REGION Network 15: EM - Abort Command
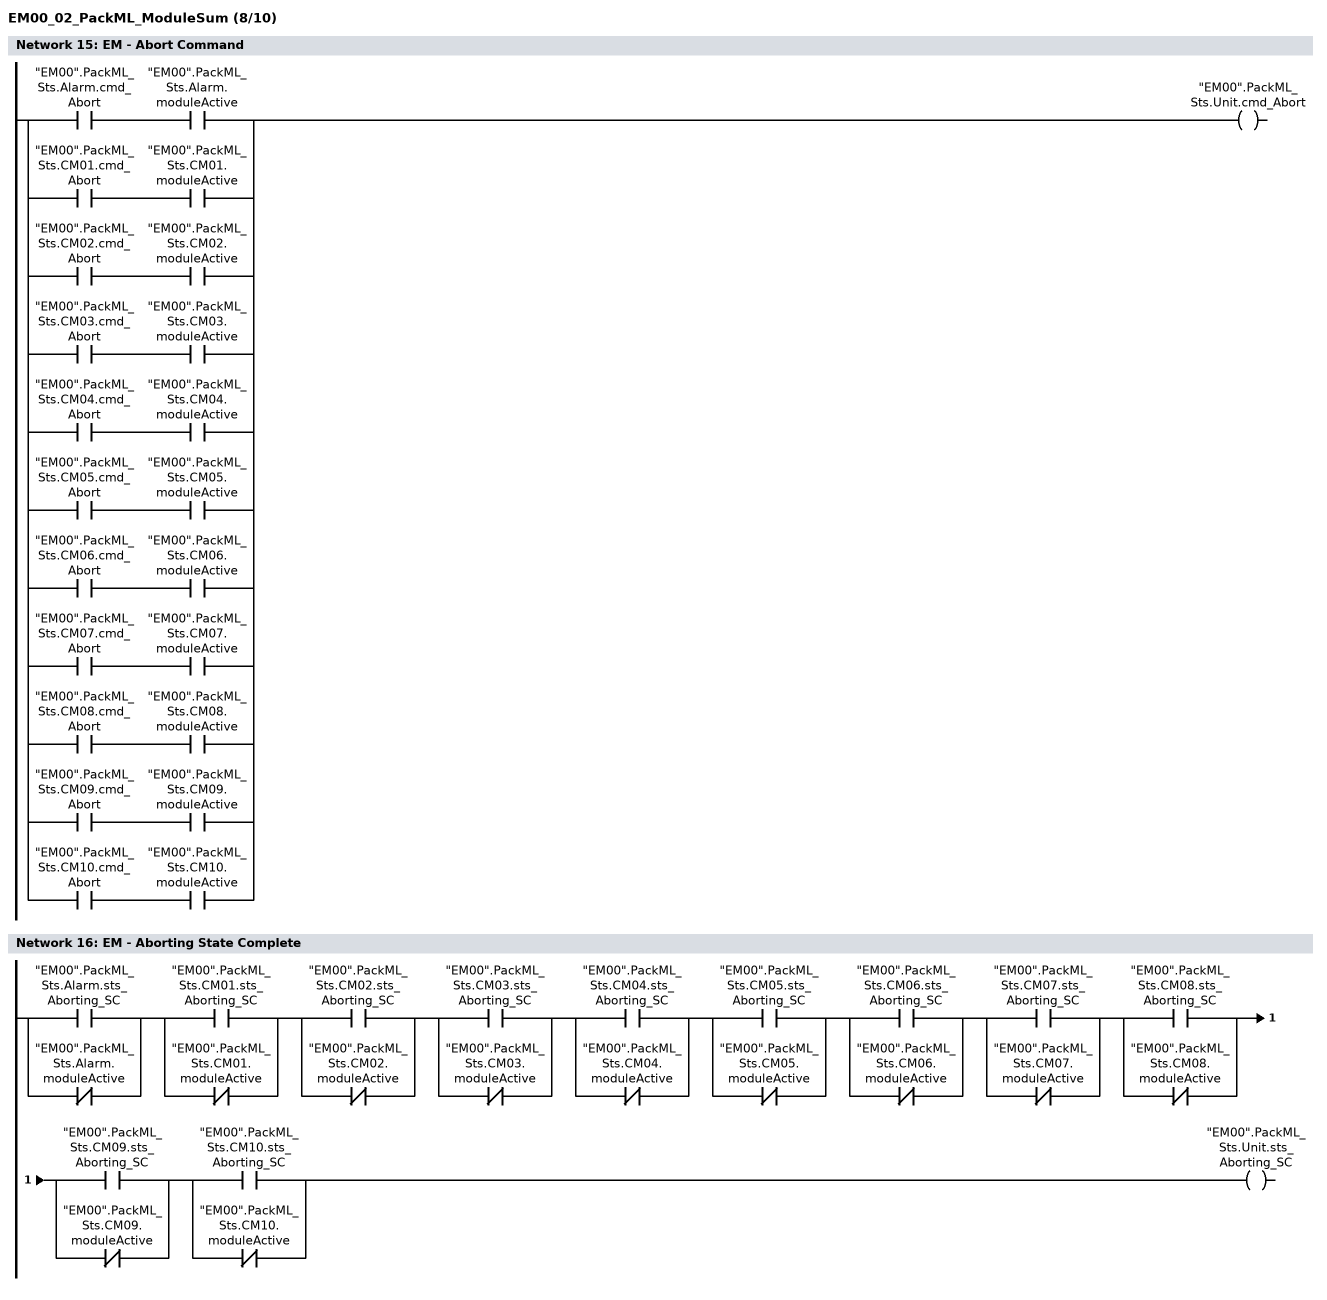
   RUNG wire#powerrail
      Contact( "EM00".PackML_Sts.Alarm.cmd_Abort )
      Contact( "EM00".PackML_Sts.Alarm.moduleActive )
      wire#w1
      Coil( "EM00".PackML_Sts.Unit.cmd_Abort )
   END_RUNG
   RUNG wire#powerrail
      Contact( "EM00".PackML_Sts.CM01.cmd_Abort )
      Contact( "EM00".PackML_Sts.CM01.moduleActive )
   END_RUNG wire#w1
   RUNG wire#powerrail
      Contact( "EM00".PackML_Sts.CM02.cmd_Abort )
      Contact( "EM00".PackML_Sts.CM02.moduleActive )
   END_RUNG wire#w1
   RUNG wire#powerrail
      Contact( "EM00".PackML_Sts.CM03.cmd_Abort )
      Contact( "EM00".PackML_Sts.CM03.moduleActive )
   END_RUNG wire#w1
   RUNG wire#powerrail
      Contact( "EM00".PackML_Sts.CM04.cmd_Abort )
      Contact( "EM00".PackML_Sts.CM04.moduleActive )
   END_RUNG wire#w1
   RUNG wire#powerrail
      Contact( "EM00".PackML_Sts.CM05.cmd_Abort )
      Contact( "EM00".PackML_Sts.CM05.moduleActive )
   END_RUNG wire#w1
   RUNG wire#powerrail
      Contact( "EM00".PackML_Sts.CM06.cmd_Abort )
      Contact( "EM00".PackML_Sts.CM06.moduleActive )
   END_RUNG wire#w1
   RUNG wire#powerrail
      Contact( "EM00".PackML_Sts.CM07.cmd_Abort )
      Contact( "EM00".PackML_Sts.CM07.moduleActive )
   END_RUNG wire#w1
   RUNG wire#powerrail
      Contact( "EM00".PackML_Sts.CM08.cmd_Abort )
      Contact( "EM00".PackML_Sts.CM08.moduleActive )
   END_RUNG wire#w1
   RUNG wire#powerrail
      Contact( "EM00".PackML_Sts.CM09.cmd_Abort )
      Contact( "EM00".PackML_Sts.CM09.moduleActive )
   END_RUNG wire#w1
   RUNG wire#powerrail
      Contact( "EM00".PackML_Sts.CM10.cmd_Abort )
      Contact( "EM00".PackML_Sts.CM10.moduleActive )
   END_RUNG wire#w1
   // the same network as SCL:
   "EM00".PackML_Sts.Unit.cmd_Abort := ("EM00".PackML_Sts.Alarm.cmd_Abort AND "EM00".PackML_Sts.Alarm.moduleActive) OR ("EM00".PackML_Sts.CM01.cmd_Abort AND "EM00".PackML_Sts.CM01.moduleActive) OR ("EM00".PackML_Sts.CM02.cmd_Abort AND "EM00".PackML_Sts.CM02.moduleActive) OR ("EM00".PackML_Sts.CM03.cmd_Abort AND "EM00".PackML_Sts.CM03.moduleActive) OR ("EM00".PackML_Sts.CM04.cmd_Abort AND "EM00".PackML_Sts.CM04.moduleActive) OR ("EM00".PackML_Sts.CM05.cmd_Abort AND "EM00".PackML_Sts.CM05.moduleActive) OR ("EM00".PackML_Sts.CM06.cmd_Abort AND "EM00".PackML_Sts.CM06.moduleActive) OR ("EM00".PackML_Sts.CM07.cmd_Abort AND "EM00".PackML_Sts.CM07.moduleActive) OR ("EM00".PackML_Sts.CM08.cmd_Abort AND "EM00".PackML_Sts.CM08.moduleActive) OR ("EM00".PackML_Sts.CM09.cmd_Abort AND "EM00".PackML_Sts.CM09.moduleActive) OR ("EM00".PackML_Sts.CM10.cmd_Abort AND "EM00".PackML_Sts.CM10.moduleActive);
END_REGION

REGION Network 16: EM - Aborting State Complete
   RUNG wire#powerrail
      Contact( "EM00".PackML_Sts.Alarm.sts_Aborting_SC )
      wire#w1
      Contact( "EM00".PackML_Sts.CM01.sts_Aborting_SC )
      wire#w2
      Contact( "EM00".PackML_Sts.CM02.sts_Aborting_SC )
      wire#w3
      Contact( "EM00".PackML_Sts.CM03.sts_Aborting_SC )
      wire#w4
      Contact( "EM00".PackML_Sts.CM04.sts_Aborting_SC )
      wire#w5
      Contact( "EM00".PackML_Sts.CM05.sts_Aborting_SC )
      wire#w6
      Contact( "EM00".PackML_Sts.CM06.sts_Aborting_SC )
      wire#w7
      Contact( "EM00".PackML_Sts.CM07.sts_Aborting_SC )
      wire#w8
      Contact( "EM00".PackML_Sts.CM08.sts_Aborting_SC )
      wire#w9
      Contact( "EM00".PackML_Sts.CM09.sts_Aborting_SC )
      wire#w10
      Contact( "EM00".PackML_Sts.CM10.sts_Aborting_SC )
      wire#w11
      Coil( "EM00".PackML_Sts.Unit.sts_Aborting_SC )
   END_RUNG
   RUNG wire#powerrail
      I_Contact( "EM00".PackML_Sts.Alarm.moduleActive )
   END_RUNG wire#w1
   RUNG wire#w1
      I_Contact( "EM00".PackML_Sts.CM01.moduleActive )
   END_RUNG wire#w2
   RUNG wire#w2
      I_Contact( "EM00".PackML_Sts.CM02.moduleActive )
   END_RUNG wire#w3
   RUNG wire#w3
      I_Contact( "EM00".PackML_Sts.CM03.moduleActive )
   END_RUNG wire#w4
   RUNG wire#w4
      I_Contact( "EM00".PackML_Sts.CM04.moduleActive )
   END_RUNG wire#w5
   RUNG wire#w5
      I_Contact( "EM00".PackML_Sts.CM05.moduleActive )
   END_RUNG wire#w6
   RUNG wire#w6
      I_Contact( "EM00".PackML_Sts.CM06.moduleActive )
   END_RUNG wire#w7
   RUNG wire#w7
      I_Contact( "EM00".PackML_Sts.CM07.moduleActive )
   END_RUNG wire#w8
   RUNG wire#w8
      I_Contact( "EM00".PackML_Sts.CM08.moduleActive )
   END_RUNG wire#w9
   RUNG wire#w9
      I_Contact( "EM00".PackML_Sts.CM09.moduleActive )
   END_RUNG wire#w10
   RUNG wire#w10
      I_Contact( "EM00".PackML_Sts.CM10.moduleActive )
   END_RUNG wire#w11
   // the same network as SCL:
   "EM00".PackML_Sts.Unit.sts_Aborting_SC := ("EM00".PackML_Sts.Alarm.sts_Aborting_SC OR NOT "EM00".PackML_Sts.Alarm.moduleActive) AND ("EM00".PackML_Sts.CM01.sts_Aborting_SC OR NOT "EM00".PackML_Sts.CM01.moduleActive) AND ("EM00".PackML_Sts.CM02.sts_Aborting_SC OR NOT "EM00".PackML_Sts.CM02.moduleActive) AND ("EM00".PackML_Sts.CM03.sts_Aborting_SC OR NOT "EM00".PackML_Sts.CM03.moduleActive) AND ("EM00".PackML_Sts.CM04.sts_Aborting_SC OR NOT "EM00".PackML_Sts.CM04.moduleActive) AND ("EM00".PackML_Sts.CM05.sts_Aborting_SC OR NOT "EM00".PackML_Sts.CM05.moduleActive) AND ("EM00".PackML_Sts.CM06.sts_Aborting_SC OR NOT "EM00".PackML_Sts.CM06.moduleActive) AND ("EM00".PackML_Sts.CM07.sts_Aborting_SC OR NOT "EM00".PackML_Sts.CM07.moduleActive) AND ("EM00".PackML_Sts.CM08.sts_Aborting_SC OR NOT "EM00".PackML_Sts.CM08.moduleActive) AND ("EM00".PackML_Sts.CM09.sts_Aborting_SC OR NOT "EM00".PackML_Sts.CM09.moduleActive) AND ("EM00".PackML_Sts.CM10.sts_Aborting_SC OR NOT "EM00".PackML_Sts.CM10.moduleActive);
END_REGION

REGION Network 17: EM - Clear Command
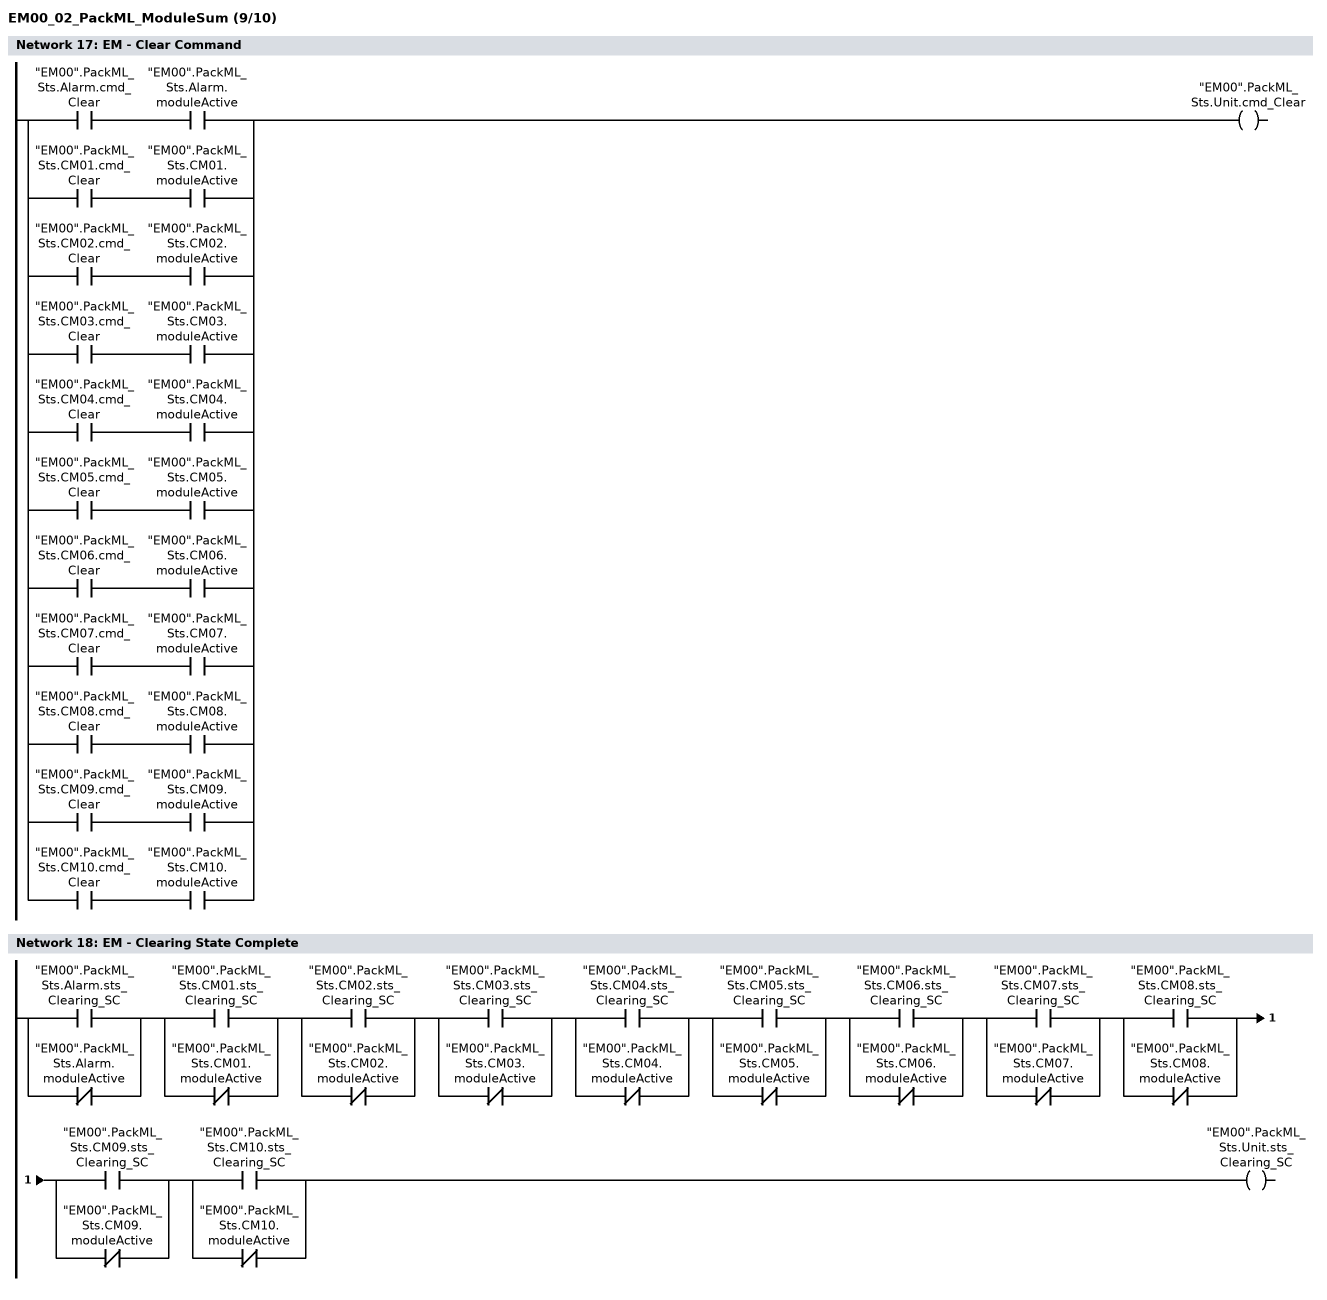
   RUNG wire#powerrail
      Contact( "EM00".PackML_Sts.Alarm.cmd_Clear )
      Contact( "EM00".PackML_Sts.Alarm.moduleActive )
      wire#w1
      Coil( "EM00".PackML_Sts.Unit.cmd_Clear )
   END_RUNG
   RUNG wire#powerrail
      Contact( "EM00".PackML_Sts.CM01.cmd_Clear )
      Contact( "EM00".PackML_Sts.CM01.moduleActive )
   END_RUNG wire#w1
   RUNG wire#powerrail
      Contact( "EM00".PackML_Sts.CM02.cmd_Clear )
      Contact( "EM00".PackML_Sts.CM02.moduleActive )
   END_RUNG wire#w1
   RUNG wire#powerrail
      Contact( "EM00".PackML_Sts.CM03.cmd_Clear )
      Contact( "EM00".PackML_Sts.CM03.moduleActive )
   END_RUNG wire#w1
   RUNG wire#powerrail
      Contact( "EM00".PackML_Sts.CM04.cmd_Clear )
      Contact( "EM00".PackML_Sts.CM04.moduleActive )
   END_RUNG wire#w1
   RUNG wire#powerrail
      Contact( "EM00".PackML_Sts.CM05.cmd_Clear )
      Contact( "EM00".PackML_Sts.CM05.moduleActive )
   END_RUNG wire#w1
   RUNG wire#powerrail
      Contact( "EM00".PackML_Sts.CM06.cmd_Clear )
      Contact( "EM00".PackML_Sts.CM06.moduleActive )
   END_RUNG wire#w1
   RUNG wire#powerrail
      Contact( "EM00".PackML_Sts.CM07.cmd_Clear )
      Contact( "EM00".PackML_Sts.CM07.moduleActive )
   END_RUNG wire#w1
   RUNG wire#powerrail
      Contact( "EM00".PackML_Sts.CM08.cmd_Clear )
      Contact( "EM00".PackML_Sts.CM08.moduleActive )
   END_RUNG wire#w1
   RUNG wire#powerrail
      Contact( "EM00".PackML_Sts.CM09.cmd_Clear )
      Contact( "EM00".PackML_Sts.CM09.moduleActive )
   END_RUNG wire#w1
   RUNG wire#powerrail
      Contact( "EM00".PackML_Sts.CM10.cmd_Clear )
      Contact( "EM00".PackML_Sts.CM10.moduleActive )
   END_RUNG wire#w1
   // the same network as SCL:
   "EM00".PackML_Sts.Unit.cmd_Clear := ("EM00".PackML_Sts.Alarm.cmd_Clear AND "EM00".PackML_Sts.Alarm.moduleActive) OR ("EM00".PackML_Sts.CM01.cmd_Clear AND "EM00".PackML_Sts.CM01.moduleActive) OR ("EM00".PackML_Sts.CM02.cmd_Clear AND "EM00".PackML_Sts.CM02.moduleActive) OR ("EM00".PackML_Sts.CM03.cmd_Clear AND "EM00".PackML_Sts.CM03.moduleActive) OR ("EM00".PackML_Sts.CM04.cmd_Clear AND "EM00".PackML_Sts.CM04.moduleActive) OR ("EM00".PackML_Sts.CM05.cmd_Clear AND "EM00".PackML_Sts.CM05.moduleActive) OR ("EM00".PackML_Sts.CM06.cmd_Clear AND "EM00".PackML_Sts.CM06.moduleActive) OR ("EM00".PackML_Sts.CM07.cmd_Clear AND "EM00".PackML_Sts.CM07.moduleActive) OR ("EM00".PackML_Sts.CM08.cmd_Clear AND "EM00".PackML_Sts.CM08.moduleActive) OR ("EM00".PackML_Sts.CM09.cmd_Clear AND "EM00".PackML_Sts.CM09.moduleActive) OR ("EM00".PackML_Sts.CM10.cmd_Clear AND "EM00".PackML_Sts.CM10.moduleActive);
END_REGION

REGION Network 18: EM - Clearing State Complete
   RUNG wire#powerrail
      Contact( "EM00".PackML_Sts.Alarm.sts_Clearing_SC )
      wire#w1
      Contact( "EM00".PackML_Sts.CM01.sts_Clearing_SC )
      wire#w2
      Contact( "EM00".PackML_Sts.CM02.sts_Clearing_SC )
      wire#w3
      Contact( "EM00".PackML_Sts.CM03.sts_Clearing_SC )
      wire#w4
      Contact( "EM00".PackML_Sts.CM04.sts_Clearing_SC )
      wire#w5
      Contact( "EM00".PackML_Sts.CM05.sts_Clearing_SC )
      wire#w6
      Contact( "EM00".PackML_Sts.CM06.sts_Clearing_SC )
      wire#w7
      Contact( "EM00".PackML_Sts.CM07.sts_Clearing_SC )
      wire#w8
      Contact( "EM00".PackML_Sts.CM08.sts_Clearing_SC )
      wire#w9
      Contact( "EM00".PackML_Sts.CM09.sts_Clearing_SC )
      wire#w10
      Contact( "EM00".PackML_Sts.CM10.sts_Clearing_SC )
      wire#w11
      Coil( "EM00".PackML_Sts.Unit.sts_Clearing_SC )
   END_RUNG
   RUNG wire#powerrail
      I_Contact( "EM00".PackML_Sts.Alarm.moduleActive )
   END_RUNG wire#w1
   RUNG wire#w1
      I_Contact( "EM00".PackML_Sts.CM01.moduleActive )
   END_RUNG wire#w2
   RUNG wire#w2
      I_Contact( "EM00".PackML_Sts.CM02.moduleActive )
   END_RUNG wire#w3
   RUNG wire#w3
      I_Contact( "EM00".PackML_Sts.CM03.moduleActive )
   END_RUNG wire#w4
   RUNG wire#w4
      I_Contact( "EM00".PackML_Sts.CM04.moduleActive )
   END_RUNG wire#w5
   RUNG wire#w5
      I_Contact( "EM00".PackML_Sts.CM05.moduleActive )
   END_RUNG wire#w6
   RUNG wire#w6
      I_Contact( "EM00".PackML_Sts.CM06.moduleActive )
   END_RUNG wire#w7
   RUNG wire#w7
      I_Contact( "EM00".PackML_Sts.CM07.moduleActive )
   END_RUNG wire#w8
   RUNG wire#w8
      I_Contact( "EM00".PackML_Sts.CM08.moduleActive )
   END_RUNG wire#w9
   RUNG wire#w9
      I_Contact( "EM00".PackML_Sts.CM09.moduleActive )
   END_RUNG wire#w10
   RUNG wire#w10
      I_Contact( "EM00".PackML_Sts.CM10.moduleActive )
   END_RUNG wire#w11
   // the same network as SCL:
   "EM00".PackML_Sts.Unit.sts_Clearing_SC := ("EM00".PackML_Sts.Alarm.sts_Clearing_SC OR NOT "EM00".PackML_Sts.Alarm.moduleActive) AND ("EM00".PackML_Sts.CM01.sts_Clearing_SC OR NOT "EM00".PackML_Sts.CM01.moduleActive) AND ("EM00".PackML_Sts.CM02.sts_Clearing_SC OR NOT "EM00".PackML_Sts.CM02.moduleActive) AND ("EM00".PackML_Sts.CM03.sts_Clearing_SC OR NOT "EM00".PackML_Sts.CM03.moduleActive) AND ("EM00".PackML_Sts.CM04.sts_Clearing_SC OR NOT "EM00".PackML_Sts.CM04.moduleActive) AND ("EM00".PackML_Sts.CM05.sts_Clearing_SC OR NOT "EM00".PackML_Sts.CM05.moduleActive) AND ("EM00".PackML_Sts.CM06.sts_Clearing_SC OR NOT "EM00".PackML_Sts.CM06.moduleActive) AND ("EM00".PackML_Sts.CM07.sts_Clearing_SC OR NOT "EM00".PackML_Sts.CM07.moduleActive) AND ("EM00".PackML_Sts.CM08.sts_Clearing_SC OR NOT "EM00".PackML_Sts.CM08.moduleActive) AND ("EM00".PackML_Sts.CM09.sts_Clearing_SC OR NOT "EM00".PackML_Sts.CM09.moduleActive) AND ("EM00".PackML_Sts.CM10.sts_Clearing_SC OR NOT "EM00".PackML_Sts.CM10.moduleActive);
END_REGION

REGION Network 19: EM - Execute State Complete
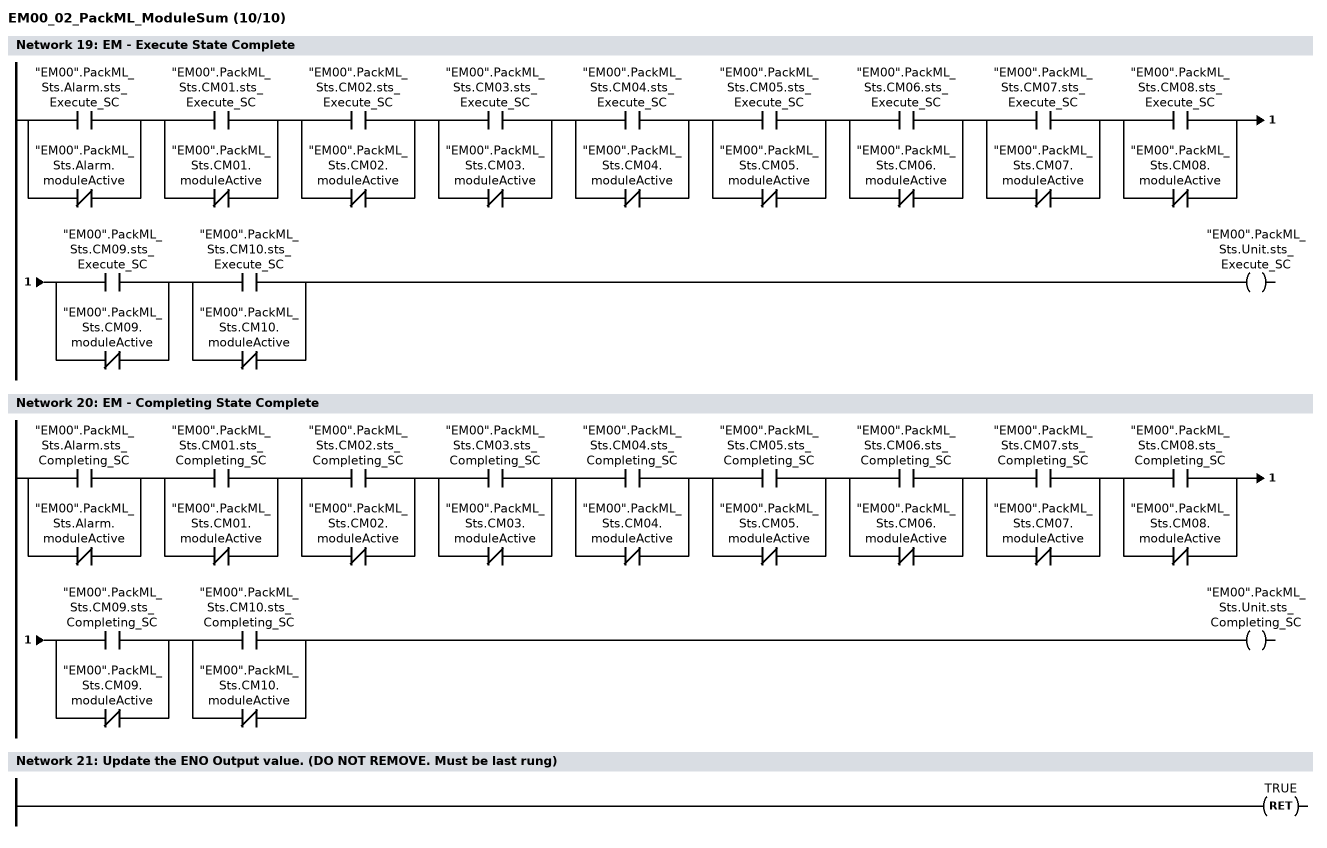
   RUNG wire#powerrail
      Contact( "EM00".PackML_Sts.Alarm.sts_Execute_SC )
      wire#w1
      Contact( "EM00".PackML_Sts.CM01.sts_Execute_SC )
      wire#w2
      Contact( "EM00".PackML_Sts.CM02.sts_Execute_SC )
      wire#w3
      Contact( "EM00".PackML_Sts.CM03.sts_Execute_SC )
      wire#w4
      Contact( "EM00".PackML_Sts.CM04.sts_Execute_SC )
      wire#w5
      Contact( "EM00".PackML_Sts.CM05.sts_Execute_SC )
      wire#w6
      Contact( "EM00".PackML_Sts.CM06.sts_Execute_SC )
      wire#w7
      Contact( "EM00".PackML_Sts.CM07.sts_Execute_SC )
      wire#w8
      Contact( "EM00".PackML_Sts.CM08.sts_Execute_SC )
      wire#w9
      Contact( "EM00".PackML_Sts.CM09.sts_Execute_SC )
      wire#w10
      Contact( "EM00".PackML_Sts.CM10.sts_Execute_SC )
      wire#w11
      Coil( "EM00".PackML_Sts.Unit.sts_Execute_SC )
   END_RUNG
   RUNG wire#powerrail
      I_Contact( "EM00".PackML_Sts.Alarm.moduleActive )
   END_RUNG wire#w1
   RUNG wire#w1
      I_Contact( "EM00".PackML_Sts.CM01.moduleActive )
   END_RUNG wire#w2
   RUNG wire#w2
      I_Contact( "EM00".PackML_Sts.CM02.moduleActive )
   END_RUNG wire#w3
   RUNG wire#w3
      I_Contact( "EM00".PackML_Sts.CM03.moduleActive )
   END_RUNG wire#w4
   RUNG wire#w4
      I_Contact( "EM00".PackML_Sts.CM04.moduleActive )
   END_RUNG wire#w5
   RUNG wire#w5
      I_Contact( "EM00".PackML_Sts.CM05.moduleActive )
   END_RUNG wire#w6
   RUNG wire#w6
      I_Contact( "EM00".PackML_Sts.CM06.moduleActive )
   END_RUNG wire#w7
   RUNG wire#w7
      I_Contact( "EM00".PackML_Sts.CM07.moduleActive )
   END_RUNG wire#w8
   RUNG wire#w8
      I_Contact( "EM00".PackML_Sts.CM08.moduleActive )
   END_RUNG wire#w9
   RUNG wire#w9
      I_Contact( "EM00".PackML_Sts.CM09.moduleActive )
   END_RUNG wire#w10
   RUNG wire#w10
      I_Contact( "EM00".PackML_Sts.CM10.moduleActive )
   END_RUNG wire#w11
   // the same network as SCL:
   "EM00".PackML_Sts.Unit.sts_Execute_SC := ("EM00".PackML_Sts.Alarm.sts_Execute_SC OR NOT "EM00".PackML_Sts.Alarm.moduleActive) AND ("EM00".PackML_Sts.CM01.sts_Execute_SC OR NOT "EM00".PackML_Sts.CM01.moduleActive) AND ("EM00".PackML_Sts.CM02.sts_Execute_SC OR NOT "EM00".PackML_Sts.CM02.moduleActive) AND ("EM00".PackML_Sts.CM03.sts_Execute_SC OR NOT "EM00".PackML_Sts.CM03.moduleActive) AND ("EM00".PackML_Sts.CM04.sts_Execute_SC OR NOT "EM00".PackML_Sts.CM04.moduleActive) AND ("EM00".PackML_Sts.CM05.sts_Execute_SC OR NOT "EM00".PackML_Sts.CM05.moduleActive) AND ("EM00".PackML_Sts.CM06.sts_Execute_SC OR NOT "EM00".PackML_Sts.CM06.moduleActive) AND ("EM00".PackML_Sts.CM07.sts_Execute_SC OR NOT "EM00".PackML_Sts.CM07.moduleActive) AND ("EM00".PackML_Sts.CM08.sts_Execute_SC OR NOT "EM00".PackML_Sts.CM08.moduleActive) AND ("EM00".PackML_Sts.CM09.sts_Execute_SC OR NOT "EM00".PackML_Sts.CM09.moduleActive) AND ("EM00".PackML_Sts.CM10.sts_Execute_SC OR NOT "EM00".PackML_Sts.CM10.moduleActive);
END_REGION

REGION Network 20: EM - Completing State Complete
   RUNG wire#powerrail
      Contact( "EM00".PackML_Sts.Alarm.sts_Completing_SC )
      wire#w1
      Contact( "EM00".PackML_Sts.CM01.sts_Completing_SC )
      wire#w2
      Contact( "EM00".PackML_Sts.CM02.sts_Completing_SC )
      wire#w3
      Contact( "EM00".PackML_Sts.CM03.sts_Completing_SC )
      wire#w4
      Contact( "EM00".PackML_Sts.CM04.sts_Completing_SC )
      wire#w5
      Contact( "EM00".PackML_Sts.CM05.sts_Completing_SC )
      wire#w6
      Contact( "EM00".PackML_Sts.CM06.sts_Completing_SC )
      wire#w7
      Contact( "EM00".PackML_Sts.CM07.sts_Completing_SC )
      wire#w8
      Contact( "EM00".PackML_Sts.CM08.sts_Completing_SC )
      wire#w9
      Contact( "EM00".PackML_Sts.CM09.sts_Completing_SC )
      wire#w10
      Contact( "EM00".PackML_Sts.CM10.sts_Completing_SC )
      wire#w11
      Coil( "EM00".PackML_Sts.Unit.sts_Completing_SC )
   END_RUNG
   RUNG wire#powerrail
      I_Contact( "EM00".PackML_Sts.Alarm.moduleActive )
   END_RUNG wire#w1
   RUNG wire#w1
      I_Contact( "EM00".PackML_Sts.CM01.moduleActive )
   END_RUNG wire#w2
   RUNG wire#w2
      I_Contact( "EM00".PackML_Sts.CM02.moduleActive )
   END_RUNG wire#w3
   RUNG wire#w3
      I_Contact( "EM00".PackML_Sts.CM03.moduleActive )
   END_RUNG wire#w4
   RUNG wire#w4
      I_Contact( "EM00".PackML_Sts.CM04.moduleActive )
   END_RUNG wire#w5
   RUNG wire#w5
      I_Contact( "EM00".PackML_Sts.CM05.moduleActive )
   END_RUNG wire#w6
   RUNG wire#w6
      I_Contact( "EM00".PackML_Sts.CM06.moduleActive )
   END_RUNG wire#w7
   RUNG wire#w7
      I_Contact( "EM00".PackML_Sts.CM07.moduleActive )
   END_RUNG wire#w8
   RUNG wire#w8
      I_Contact( "EM00".PackML_Sts.CM08.moduleActive )
   END_RUNG wire#w9
   RUNG wire#w9
      I_Contact( "EM00".PackML_Sts.CM09.moduleActive )
   END_RUNG wire#w10
   RUNG wire#w10
      I_Contact( "EM00".PackML_Sts.CM10.moduleActive )
   END_RUNG wire#w11
   // the same network as SCL:
   "EM00".PackML_Sts.Unit.sts_Completing_SC := ("EM00".PackML_Sts.Alarm.sts_Completing_SC OR NOT "EM00".PackML_Sts.Alarm.moduleActive) AND ("EM00".PackML_Sts.CM01.sts_Completing_SC OR NOT "EM00".PackML_Sts.CM01.moduleActive) AND ("EM00".PackML_Sts.CM02.sts_Completing_SC OR NOT "EM00".PackML_Sts.CM02.moduleActive) AND ("EM00".PackML_Sts.CM03.sts_Completing_SC OR NOT "EM00".PackML_Sts.CM03.moduleActive) AND ("EM00".PackML_Sts.CM04.sts_Completing_SC OR NOT "EM00".PackML_Sts.CM04.moduleActive) AND ("EM00".PackML_Sts.CM05.sts_Completing_SC OR NOT "EM00".PackML_Sts.CM05.moduleActive) AND ("EM00".PackML_Sts.CM06.sts_Completing_SC OR NOT "EM00".PackML_Sts.CM06.moduleActive) AND ("EM00".PackML_Sts.CM07.sts_Completing_SC OR NOT "EM00".PackML_Sts.CM07.moduleActive) AND ("EM00".PackML_Sts.CM08.sts_Completing_SC OR NOT "EM00".PackML_Sts.CM08.moduleActive) AND ("EM00".PackML_Sts.CM09.sts_Completing_SC OR NOT "EM00".PackML_Sts.CM09.moduleActive) AND ("EM00".PackML_Sts.CM10.sts_Completing_SC OR NOT "EM00".PackML_Sts.CM10.moduleActive);
END_REGION

REGION Network 21: Update the ENO Output value. (DO NOT REMOVE. Must be last rung)
   RUNG wire#powerrail
      ReturnCoil( TRUE )
   END_RUNG
   // the same network as SCL:
   ENO := TRUE;
   RETURN;
END_REGION
END_FUNCTION_BLOCK

FUNCTION_BLOCK "EM00_CM01_MainOpStation"   // FB31651, LAD
TITLE = EM00_CM01_MainOpStation
{ S7_Optimized_Access := 'TRUE' }
AUTHOR : tech.team.motioncontrol@siemens.com
FAMILY : CPG
VERSION : 1.1
// Support: tech.team.motioncontrol@siemens.com
   VAR
      instAlarm_EStop : "CPG_Event";   // Alarm Event - EStop pressed (Event instance)
      instAlarm_HMI_StopPB : "CPG_Event";   // Alarm Event - HMI Stop PB pressed (Event instance)
      instStatus_WaitingForStartCmd : "CPG_Event";   // Status Event - waiting for start command (Event instance)
      instStatus_WaitingForResetCmd : "CPG_Event";   // Status Event - waiting for reset command (Event instance)
      instAlarm_Hold_PB : "CPG_Event";   // Alarm Event - HMI Held PB pressed (Event instance)
      instStatus_WaitingForUnHoldCmd : "CPG_Event";   // Status Event - waiting for unhold command (Event instance)
      instTimer_StartingDelay_SC : IEC_TIMER;   // IEC Timer - starting delay (demo only - used to slow state model transition)
      instTimer_CompletingDelay_SC : IEC_TIMER;   // IEC Timer - completing delay (demo only - used to slow state model transition)
      instTimer_AbortingDelay_SC : IEC_TIMER;   // IEC Timer - aborting delay (demo only - used to slow state model transition)
      instTimer_StoppingDelay_SC : IEC_TIMER;   // IEC Timer - stopping delay (demo only - used to slow state model transition)
      instTimer_ResettingDelay_SC : IEC_TIMER;   // IEC Timer - resetting delay (demo only - used to slow state model transition)
      instTimer_HoldingDelay_SC : IEC_TIMER;   // IEC Timer - holding delay (demo only - used to slow state model transition)
      instTimer_UnHoldingDelay_SC : IEC_TIMER;   // IEC Timer - un-holding delay (demo only - used to slow state model transition)
      instTimer_SuspendingDelay_SC : IEC_TIMER;   // IEC Timer - suspending delay (demo only - used to slow state model transition)
      instTimer_UnSuspendingDelay_SC : IEC_TIMER;   // IEC Timer - un-suspending delay (demo only - used to slow state model transition)
      instTimer_ClearingDelay_SC : IEC_TIMER;   // IEC Timer - clearing delay (demo only - used to slow state model transition)
      FTriggerTest_Instance : "FTriggerTest";
   END_VAR
BEGIN

REGION Network 1: *** Begin the Setpoint Management Information Section ***
END_REGION

REGION Network 2: *** Begin the Logic Section ***
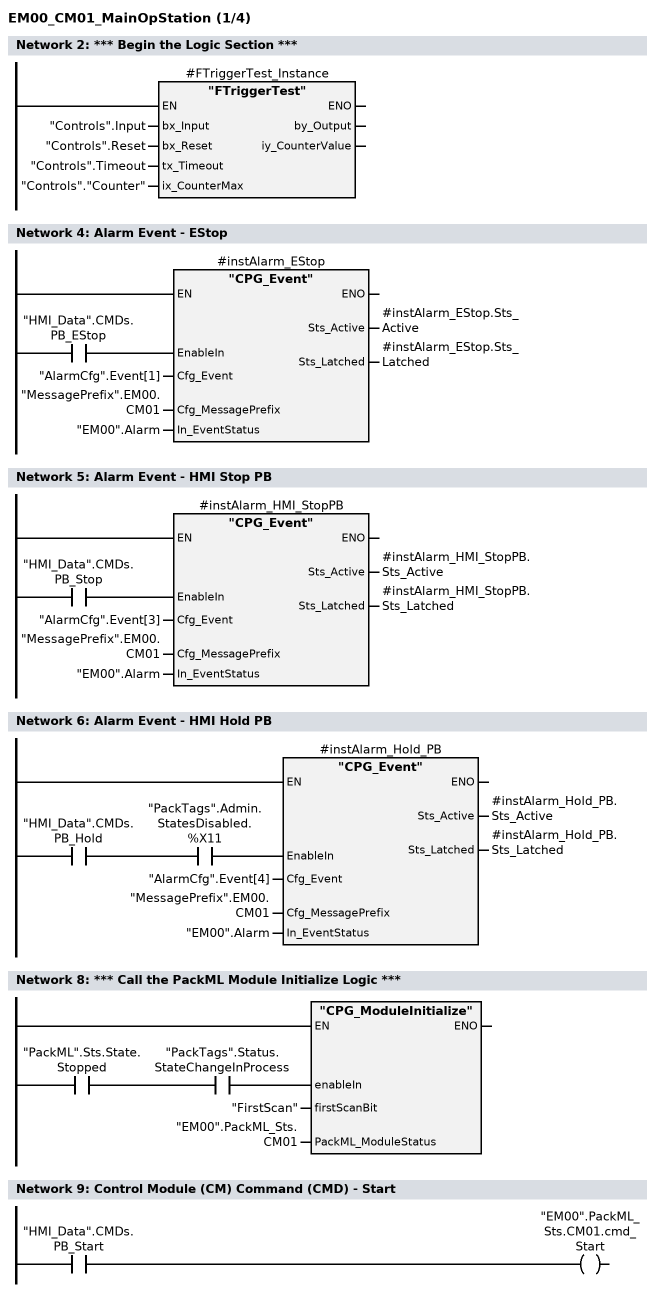
   RUNG wire#powerrail
      #FTriggerTest_Instance(bx_Input := "Controls".Input, bx_Reset := "Controls".Reset, tx_Timeout := "Controls".Timeout, ix_CounterMax := "Controls"."Counter", by_Output =>, iy_CounterValue =>)
   END_RUNG
   // the same network as SCL:
   #FTriggerTest_Instance(bx_Input := "Controls".Input,   // "FTriggerTest"
                          bx_Reset := "Controls".Reset,
                          tx_Timeout := "Controls".Timeout,
                          ix_CounterMax := "Controls"."Counter");
END_REGION

REGION Network 3: *** Begin the Event Information Section ***
END_REGION

REGION Network 4: Alarm Event - EStop
   RUNG wire#powerrail
      #instAlarm_EStop(EnableIn := wire#w1, Cfg_Event := "AlarmCfg".Event[1], Cfg_MessagePrefix := "MessagePrefix".EM00.CM01, In_EventStatus := "EM00".Alarm, Sts_Active => #instAlarm_EStop.Sts_Active, Sts_Latched => #instAlarm_EStop.Sts_Latched)
   END_RUNG
   RUNG wire#powerrail
      Contact( "HMI_Data".CMDs.PB_EStop )
   END_RUNG wire#w1
   // the same network as SCL:
   #instAlarm_EStop(EnableIn := "HMI_Data".CMDs.PB_EStop,   // "CPG_Event"
                    Cfg_Event := "AlarmCfg".Event[1],
                    Cfg_MessagePrefix := "MessagePrefix".EM00.CM01,
                    In_EventStatus := "EM00".Alarm,
                    Sts_Active => #instAlarm_EStop.Sts_Active,
                    Sts_Latched => #instAlarm_EStop.Sts_Latched);
END_REGION

REGION Network 5: Alarm Event - HMI Stop PB
   RUNG wire#powerrail
      #instAlarm_HMI_StopPB(EnableIn := wire#w1, Cfg_Event := "AlarmCfg".Event[3], Cfg_MessagePrefix := "MessagePrefix".EM00.CM01, In_EventStatus := "EM00".Alarm, Sts_Active => #instAlarm_HMI_StopPB.Sts_Active, Sts_Latched => #instAlarm_HMI_StopPB.Sts_Latched)
   END_RUNG
   RUNG wire#powerrail
      Contact( "HMI_Data".CMDs.PB_Stop )
   END_RUNG wire#w1
   // the same network as SCL:
   #instAlarm_HMI_StopPB(EnableIn := "HMI_Data".CMDs.PB_Stop,   // "CPG_Event"
                         Cfg_Event := "AlarmCfg".Event[3],
                         Cfg_MessagePrefix := "MessagePrefix".EM00.CM01,
                         In_EventStatus := "EM00".Alarm,
                         Sts_Active => #instAlarm_HMI_StopPB.Sts_Active,
                         Sts_Latched => #instAlarm_HMI_StopPB.Sts_Latched);
END_REGION

REGION Network 6: Alarm Event - HMI Hold PB
   RUNG wire#powerrail
      #instAlarm_Hold_PB(EnableIn := wire#w1, Cfg_Event := "AlarmCfg".Event[4], Cfg_MessagePrefix := "MessagePrefix".EM00.CM01, In_EventStatus := "EM00".Alarm, Sts_Active => #instAlarm_Hold_PB.Sts_Active, Sts_Latched => #instAlarm_Hold_PB.Sts_Latched)
   END_RUNG
   RUNG wire#powerrail
      Contact( "HMI_Data".CMDs.PB_Hold )
      Contact( "PackTags".Admin.StatesDisabled.%X11 )
   END_RUNG wire#w1
   // the same network as SCL:
   #instAlarm_Hold_PB(EnableIn := "HMI_Data".CMDs.PB_Hold AND "PackTags".Admin.StatesDisabled.%X11,   // "CPG_Event"
                      Cfg_Event := "AlarmCfg".Event[4],
                      Cfg_MessagePrefix := "MessagePrefix".EM00.CM01,
                      In_EventStatus := "EM00".Alarm,
                      Sts_Active => #instAlarm_Hold_PB.Sts_Active,
                      Sts_Latched => #instAlarm_Hold_PB.Sts_Latched);
END_REGION

REGION Network 7: *** Begin the State Model Status Feedback Section ***
END_REGION

REGION Network 8: *** Call the PackML Module Initialize Logic ***
   RUNG wire#powerrail
      "CPG_ModuleInitialize"(enableIn := wire#w1, firstScanBit := "FirstScan", PackML_ModuleStatus := "EM00".PackML_Sts.CM01)
   END_RUNG
   RUNG wire#powerrail
      Contact( "PackML".Sts.State.Stopped )
      Contact( "PackTags".Status.StateChangeInProcess )
   END_RUNG wire#w1
   // the same network as SCL:
   "CPG_ModuleInitialize"(enableIn := "PackML".Sts.State.Stopped AND "PackTags".Status.StateChangeInProcess,
                          firstScanBit := "FirstScan",
                          PackML_ModuleStatus := "EM00".PackML_Sts.CM01);
END_REGION

REGION Network 9: Control Module (CM) Command (CMD) - Start
   RUNG wire#powerrail
      Contact( "HMI_Data".CMDs.PB_Start )
      Coil( "EM00".PackML_Sts.CM01.cmd_Start )
   END_RUNG
   // the same network as SCL:
   "EM00".PackML_Sts.CM01.cmd_Start := "HMI_Data".CMDs.PB_Start;
END_REGION

REGION Network 10: Status Event message for HMI - Waiting for Start PB
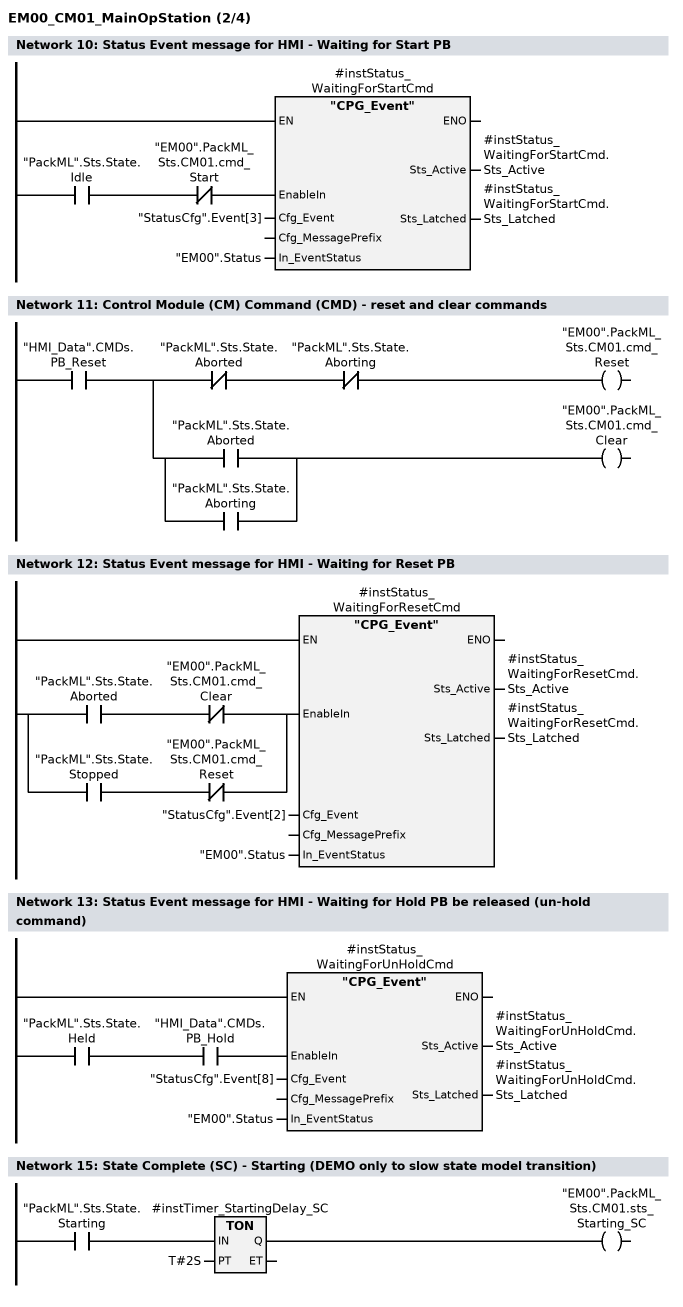
   RUNG wire#powerrail
      #instStatus_WaitingForStartCmd(EnableIn := wire#w1, Cfg_Event := "StatusCfg".Event[3], Cfg_MessagePrefix :=, In_EventStatus := "EM00".Status, Sts_Active => #instStatus_WaitingForStartCmd.Sts_Active, Sts_Latched => #instStatus_WaitingForStartCmd.Sts_Latched)
   END_RUNG
   RUNG wire#powerrail
      Contact( "PackML".Sts.State.Idle )
      I_Contact( "EM00".PackML_Sts.CM01.cmd_Start )
   END_RUNG wire#w1
   // the same network as SCL:
   #instStatus_WaitingForStartCmd(EnableIn := "PackML".Sts.State.Idle AND NOT "EM00".PackML_Sts.CM01.cmd_Start,   // "CPG_Event"
                           Cfg_Event := "StatusCfg".Event[3],
                           In_EventStatus := "EM00".Status,
                           Sts_Active => #instStatus_WaitingForStartCmd.Sts_Active,
                           Sts_Latched => #instStatus_WaitingForStartCmd.Sts_Latched);
END_REGION

REGION Network 11: Control Module (CM) Command (CMD) - reset and clear commands
   RUNG wire#powerrail
      Contact( "HMI_Data".CMDs.PB_Reset )
      wire#w1
      I_Contact( "PackML".Sts.State.Aborted )
      I_Contact( "PackML".Sts.State.Aborting )
      Coil( "EM00".PackML_Sts.CM01.cmd_Reset )
   END_RUNG
   RUNG wire#w1
      Contact( "PackML".Sts.State.Aborted )
      wire#w2
      Coil( "EM00".PackML_Sts.CM01.cmd_Clear )
   END_RUNG
   RUNG wire#w1
      Contact( "PackML".Sts.State.Aborting )
   END_RUNG wire#w2
   // the same network as SCL:
   "EM00".PackML_Sts.CM01.cmd_Reset := "HMI_Data".CMDs.PB_Reset AND NOT "PackML".Sts.State.Aborted AND NOT "PackML".Sts.State.Aborting;
   "EM00".PackML_Sts.CM01.cmd_Clear := "HMI_Data".CMDs.PB_Reset AND ("PackML".Sts.State.Aborted OR "PackML".Sts.State.Aborting);
END_REGION

REGION Network 12: Status Event message for HMI - Waiting for Reset PB
   RUNG wire#powerrail
      #instStatus_WaitingForResetCmd(EnableIn := wire#w1, Cfg_Event := "StatusCfg".Event[2], Cfg_MessagePrefix :=, In_EventStatus := "EM00".Status, Sts_Active => #instStatus_WaitingForResetCmd.Sts_Active, Sts_Latched => #instStatus_WaitingForResetCmd.Sts_Latched)
   END_RUNG
   RUNG wire#powerrail
      Contact( "PackML".Sts.State.Aborted )
      I_Contact( "EM00".PackML_Sts.CM01.cmd_Clear )
   END_RUNG wire#w1
   RUNG wire#powerrail
      Contact( "PackML".Sts.State.Stopped )
      I_Contact( "EM00".PackML_Sts.CM01.cmd_Reset )
   END_RUNG wire#w1
   // the same network as SCL:
   #instStatus_WaitingForResetCmd(EnableIn := ("PackML".Sts.State.Aborted AND NOT "EM00".PackML_Sts.CM01.cmd_Clear) OR ("PackML".Sts.State.Stopped AND NOT "EM00".PackML_Sts.CM01.cmd_Reset),   // "CPG_Event"
                           Cfg_Event := "StatusCfg".Event[2],
                           In_EventStatus := "EM00".Status,
                           Sts_Active => #instStatus_WaitingForResetCmd.Sts_Active,
                           Sts_Latched => #instStatus_WaitingForResetCmd.Sts_Latched);
END_REGION

REGION Network 13: Status Event message for HMI - Waiting for Hold PB be released (un-hold command)
   RUNG wire#powerrail
      #instStatus_WaitingForUnHoldCmd(EnableIn := wire#w1, Cfg_Event := "StatusCfg".Event[8], Cfg_MessagePrefix :=, In_EventStatus := "EM00".Status, Sts_Active => #instStatus_WaitingForUnHoldCmd.Sts_Active, Sts_Latched => #instStatus_WaitingForUnHoldCmd.Sts_Latched)
   END_RUNG
   RUNG wire#powerrail
      Contact( "PackML".Sts.State.Held )
      Contact( "HMI_Data".CMDs.PB_Hold )
   END_RUNG wire#w1
   // the same network as SCL:
   #instStatus_WaitingForUnHoldCmd(EnableIn := "PackML".Sts.State.Held AND "HMI_Data".CMDs.PB_Hold,   // "CPG_Event"
                           Cfg_Event := "StatusCfg".Event[8],
                           In_EventStatus := "EM00".Status,
                           Sts_Active => #instStatus_WaitingForUnHoldCmd.Sts_Active,
                           Sts_Latched => #instStatus_WaitingForUnHoldCmd.Sts_Latched);
END_REGION

REGION Network 14: State Model delay timers used to slow state model transition - only used for demo purposes (remove for real projects)
END_REGION

REGION Network 15: State Complete (SC) - Starting (DEMO only to slow state model transition)
   #instTimer_StartingDelay_SC.TON(IN := "PackML".Sts.State.Starting, PT := T#2S);
   "EM00".PackML_Sts.CM01.sts_Starting_SC := #instTimer_StartingDelay_SC.Q;
END_REGION

REGION Network 16: State Complete (SC) - Completing (DEMO only to slow state model transition)
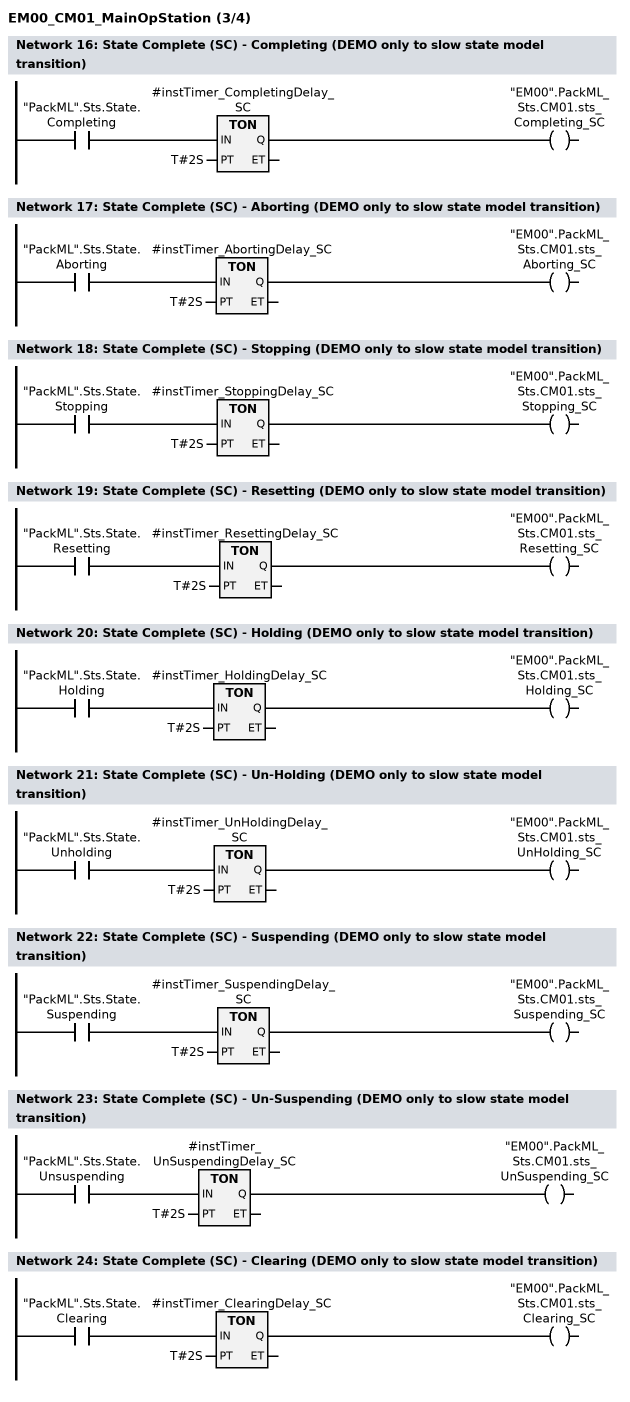
   #instTimer_CompletingDelay_SC.TON(IN := "PackML".Sts.State.Completing, PT := T#2S);
   "EM00".PackML_Sts.CM01.sts_Completing_SC := #instTimer_CompletingDelay_SC.Q;
END_REGION

REGION Network 17: State Complete (SC) - Aborting (DEMO only to slow state model transition)
   #instTimer_AbortingDelay_SC.TON(IN := "PackML".Sts.State.Aborting, PT := T#2S);
   "EM00".PackML_Sts.CM01.sts_Aborting_SC := #instTimer_AbortingDelay_SC.Q;
END_REGION

REGION Network 18: State Complete (SC) - Stopping (DEMO only to slow state model transition)
   #instTimer_StoppingDelay_SC.TON(IN := "PackML".Sts.State.Stopping, PT := T#2S);
   "EM00".PackML_Sts.CM01.sts_Stopping_SC := #instTimer_StoppingDelay_SC.Q;
END_REGION

REGION Network 19: State Complete (SC) - Resetting (DEMO only to slow state model transition)
   #instTimer_ResettingDelay_SC.TON(IN := "PackML".Sts.State.Resetting, PT := T#2S);
   "EM00".PackML_Sts.CM01.sts_Resetting_SC := #instTimer_ResettingDelay_SC.Q;
END_REGION

REGION Network 20: State Complete (SC) - Holding (DEMO only to slow state model transition)
   #instTimer_HoldingDelay_SC.TON(IN := "PackML".Sts.State.Holding, PT := T#2S);
   "EM00".PackML_Sts.CM01.sts_Holding_SC := #instTimer_HoldingDelay_SC.Q;
END_REGION

REGION Network 21: State Complete (SC) - Un-Holding (DEMO only to slow state model transition)
   #instTimer_UnHoldingDelay_SC.TON(IN := "PackML".Sts.State.Unholding, PT := T#2S);
   "EM00".PackML_Sts.CM01.sts_UnHolding_SC := #instTimer_UnHoldingDelay_SC.Q;
END_REGION

REGION Network 22: State Complete (SC) - Suspending (DEMO only to slow state model transition)
   #instTimer_SuspendingDelay_SC.TON(IN := "PackML".Sts.State.Suspending, PT := T#2S);
   "EM00".PackML_Sts.CM01.sts_Suspending_SC := #instTimer_SuspendingDelay_SC.Q;
END_REGION

REGION Network 23: State Complete (SC) - Un-Suspending (DEMO only to slow state model transition)
   #instTimer_UnSuspendingDelay_SC.TON(IN := "PackML".Sts.State.Unsuspending, PT := T#2S);
   "EM00".PackML_Sts.CM01.sts_UnSuspending_SC := #instTimer_UnSuspendingDelay_SC.Q;
END_REGION

REGION Network 24: State Complete (SC) - Clearing (DEMO only to slow state model transition)
   #instTimer_ClearingDelay_SC.TON(IN := "PackML".Sts.State.Clearing, PT := T#2S);
   "EM00".PackML_Sts.CM01.sts_Clearing_SC := #instTimer_ClearingDelay_SC.Q;
END_REGION

REGION Network 25: State Complete (SC) - Execute
   // triggering this bit will make the transition to the completing state
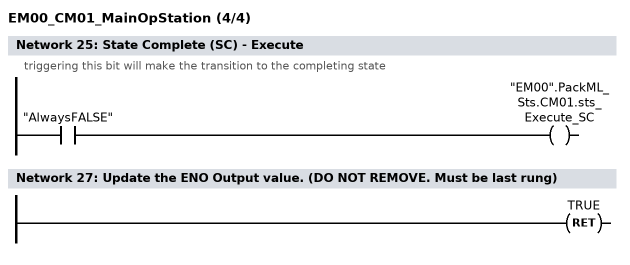
   RUNG wire#powerrail
      Contact( "AlwaysFALSE" )
      Coil( "EM00".PackML_Sts.CM01.sts_Execute_SC )
   END_RUNG
   // the same network as SCL:
   "EM00".PackML_Sts.CM01.sts_Execute_SC := "AlwaysFALSE";
END_REGION

REGION Network 27: Update the ENO Output value. (DO NOT REMOVE. Must be last rung)
   RUNG wire#powerrail
      ReturnCoil( TRUE )
   END_RUNG
   // the same network as SCL:
   ENO := TRUE;
   RETURN;
END_REGION
END_FUNCTION_BLOCK

FUNCTION_BLOCK "EM00_CM02_Conveyor"   // FB31652, LAD
TITLE = EM00_CM02_HornBeacons
{ S7_Optimized_Access := 'TRUE' }
AUTHOR : tech.team.motioncontrol@siemens.com
FAMILY : CPG
VERSION : 1.1
// Support: tech.team.motioncontrol@siemens.com
   VAR
      statDummy : Bool;   // Variable to control a horn
      instConveyor : "Conveyor";
   END_VAR
BEGIN

REGION Network 1: *** Begin the Setpoint Management Information Section ***
END_REGION

REGION Network 2: *** Begin the Logic Section ***
END_REGION

REGION Network 3: Conveyor instance